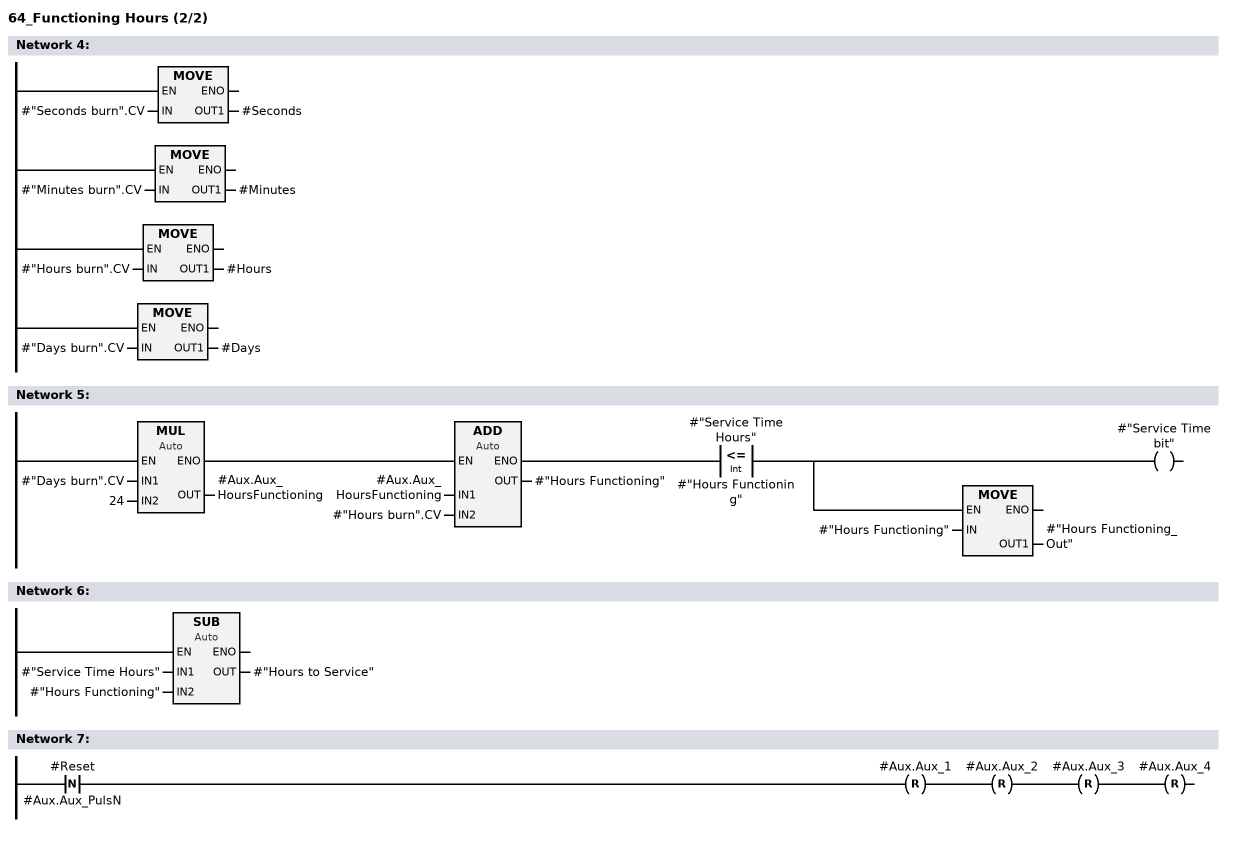
   RUNG wire#powerrail
      Move(in := #"Seconds burn".CV, out1 => #Seconds)
   END_RUNG
   RUNG wire#powerrail
      Move(in := #"Minutes burn".CV, out1 => #Minutes)
   END_RUNG
   RUNG wire#powerrail
      Move(in := #"Hours burn".CV, out1 => #Hours)
   END_RUNG
   RUNG wire#powerrail
      Move(in := #"Days burn".CV, out1 => #Days)
   END_RUNG
   // the same network as SCL:
   #Seconds := #"Seconds burn".CV;
   #Minutes := #"Minutes burn".CV;
   #Hours := #"Hours burn".CV;
   #Days := #"Days burn".CV;
END_REGION

REGION Network 5
   RUNG wire#powerrail
      Mul(in1 := #"Days burn".CV, in2 := 24, out => #Aux.Aux_HoursFunctioning)
      Add(in1 := #Aux.Aux_HoursFunctioning, in2 := #"Hours burn".CV, out => #"Hours Functioning")
      { S7_Templates := "SrcType := Int" } LE_Contact(in1 := #"Service Time Hours", in2 := #"Hours Functioning")
      wire#w1
      Coil( #"Service Time bit" )
   END_RUNG
   RUNG wire#w1
      Move(in := #"Hours Functioning", out1 => #"Hours Functioning_Out")
   END_RUNG
   // the same network as SCL:
   #Aux.Aux_HoursFunctioning := #"Days burn".CV * 24;
   #"Hours Functioning" := #Aux.Aux_HoursFunctioning + #"Hours burn".CV;
   #"Service Time bit" := #"Service Time Hours" <= #"Hours Functioning";
   IF #"Service Time bit" THEN #"Hours Functioning_Out" := #"Hours Functioning"; END_IF;
END_REGION

REGION Network 6
   RUNG wire#powerrail
      Sub(in1 := #"Service Time Hours", in2 := #"Hours Functioning", out => #"Hours to Service")
   END_RUNG
   // the same network as SCL:
   #"Hours to Service" := #"Service Time Hours" - #"Hours Functioning";
END_REGION

REGION Network 7
   RUNG wire#powerrail
      N_Contact(operand := #Reset, bit := #Aux.Aux_PulsN)
      R_Coil( #Aux.Aux_1 )
      R_Coil( #Aux.Aux_2 )
      R_Coil( #Aux.Aux_3 )
      R_Coil( #Aux.Aux_4 )
   END_RUNG
   // the same network as SCL:
   #_w1 := NOT #Reset AND #Aux.Aux_PulsN;   // falling edge of #Reset
   #Aux.Aux_PulsN := #Reset;
   IF #_w1 THEN
       #Aux.Aux_1 := FALSE;
       #Aux.Aux_2 := FALSE;
       #Aux.Aux_3 := FALSE;
       #Aux.Aux_4 := FALSE;
   END_IF;
END_REGION
END_FUNCTION_BLOCK

FUNCTION_BLOCK "503_ALARM CHCK II"   // FB507, LAD
{ S7_Optimized_Access := 'TRUE' }
VERSION : 0.1
   VAR_INPUT
      "Alarm Word 1" : Word;
      "Alarm Word Ack 1" : Word;
      "Alarm Word 2" : Word;
      "Alarm Word Ack 2" : Word;
      "Alarm Word 3" : Word;
      "Alarm Word Ack 3" : Word;
      "Alarm Word 4" : Word;
      "Alarm Word Ack 4" : Word;
      "Alarm Word 5" : Word;
      "Alarm Word Ack 5" : Word;
      "Alarm Word 6" : Word;
      "Alarm Word Ack 6" : Word;
      "Alarm Word 7" : Word;
      "Alarm Word Ack 7" : Word;
      "Alarm Word 8" : Word;
      "Alarm Word Ack 8" : Word;
      "Alarm Word 9" : Word;
      "Alarm Word 10" : Word;
      "Alarm Word 11" : Word;
      "Alarm Word 12" : Word;
      "Alarm Word 13" : Word;
      "Alarm Word 14" : Word;
      "Alarm Word 15" : Word;
      "Alarm Word 16" : Word;
      "Ack frequency" : Time;
      "Reset Alarm" : Bool;
   END_VAR
   VAR_OUTPUT
      Alarm : Bool;
      "New Alarm" : Bool;
      "Acknowledged Alarm" : Bool;
      Buzzer : Bool;
   END_VAR
   VAR
      "Alarm Word Interm 1" : Word;
      "Alarm Word Interm 2" : Word;
      "Alarm Word Interm 3" : Word;
      "Alarm Word Interm 4" : Word;
      "Alarm Word Interm 5" : Word;
      "Alarm Word Interm 6" : Word;
      "Alarm Word Interm 7" : Word;
      "Alarm Word Interm 8" : Word;
      "Alarm Word Interm 9" : Word;
      "Alarm Word Interm 10" : Word;
      "Alarm Word Interm 11" : Word;
      "Alarm Word Interm 12" : Word;
      "Alarm Word Interm 13" : Word;
      "Alarm Word Interm 14" : Word;
      "Alarm Word Interm 15" : Word;
      "Alarm Word Interm 16" : Word;
      "Alarm Word bool 1" : Bool;
      "Alarm Word bool 2" : Bool;
      "Alarm Word bool 3" : Bool;
      "Alarm Word bool 4" : Bool;
      "Alarm Word bool 5" : Bool;
      "Alarm Word bool 6" : Bool;
      "Alarm Word bool 7" : Bool;
      "Alarm Word bool 8" : Bool;
      "Alarm Word bool 9" : Bool;
      "Alarm Word bool 10" : Bool;
      "Alarm Word bool 11" : Bool;
      "Alarm Word bool 12" : Bool;
      "Alarm Word bool 13" : Bool;
      "Alarm Word bool 14" : Bool;
      "Alarm Word bool 15" : Bool;
      "Alarm Word bool 16" : Bool;
      True : Bool;
      False : Bool;
      "Delayed Alarm Reset" : TON_TIME;
      "Sound Alarm Delayed" : Bool;
      "SET TON" : TON_TIME;
      "RESET TON" : TON_TIME;
   END_VAR
   VAR_TEMP   // added for the SCL form of the ladder/FBD networks
      _w1 : Bool;
   END_VAR
BEGIN

REGION Network 1: True/False
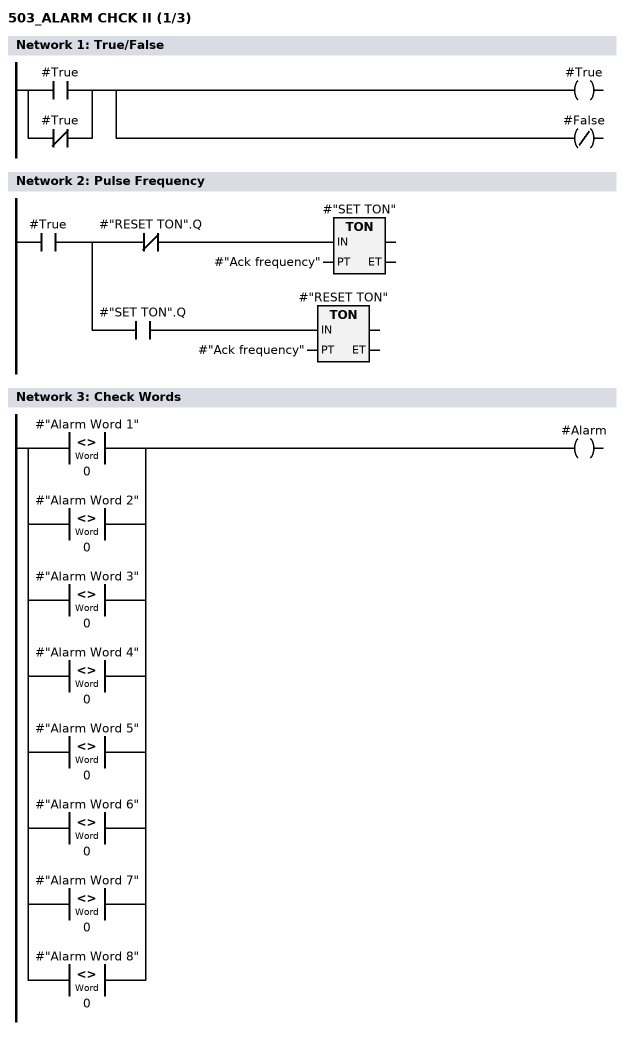
   RUNG wire#powerrail
      Contact( #True )
      wire#w1
      Coil( #True )
   END_RUNG
   RUNG wire#powerrail
      I_Contact( #True )
   END_RUNG wire#w1
   RUNG wire#w1
      I_Coil( #False )
   END_RUNG
   // the same network as SCL:
   #True := #True OR NOT #True;
   #False := NOT #True;
END_REGION

REGION Network 2: Pulse Frequency
   #"SET TON"(IN := #True AND NOT #"RESET TON".Q, PT := #"Ack frequency");   // TON
   #"RESET TON"(IN := #True AND #"SET TON".Q, PT := #"Ack frequency");   // TON
END_REGION

REGION Network 3: Check Words
   RUNG wire#powerrail
      { S7_Templates := "SrcType := Word" } NE_Contact(in1 := #"Alarm Word 1", in2 := 0)
      wire#w1
      Coil( #Alarm )
   END_RUNG
   RUNG wire#powerrail
      { S7_Templates := "SrcType := Word" } NE_Contact(in1 := #"Alarm Word 2", in2 := 0)
   END_RUNG wire#w1
   RUNG wire#powerrail
      { S7_Templates := "SrcType := Word" } NE_Contact(in1 := #"Alarm Word 3", in2 := 0)
   END_RUNG wire#w1
   RUNG wire#powerrail
      { S7_Templates := "SrcType := Word" } NE_Contact(in1 := #"Alarm Word 4", in2 := 0)
   END_RUNG wire#w1
   RUNG wire#powerrail
      { S7_Templates := "SrcType := Word" } NE_Contact(in1 := #"Alarm Word 5", in2 := 0)
   END_RUNG wire#w1
   RUNG wire#powerrail
      { S7_Templates := "SrcType := Word" } NE_Contact(in1 := #"Alarm Word 6", in2 := 0)
   END_RUNG wire#w1
   RUNG wire#powerrail
      { S7_Templates := "SrcType := Word" } NE_Contact(in1 := #"Alarm Word 7", in2 := 0)
   END_RUNG wire#w1
   RUNG wire#powerrail
      { S7_Templates := "SrcType := Word" } NE_Contact(in1 := #"Alarm Word 8", in2 := 0)
   END_RUNG wire#w1
   // the same network as SCL:
   #Alarm := (#"Alarm Word 1" <> 0) OR (#"Alarm Word 2" <> 0) OR (#"Alarm Word 3" <> 0) OR (#"Alarm Word 4" <> 0) OR (#"Alarm Word 5" <> 0) OR (#"Alarm Word 6" <> 0) OR (#"Alarm Word 7" <> 0) OR (#"Alarm Word 8" <> 0);
END_REGION

REGION Network 4: Check Words
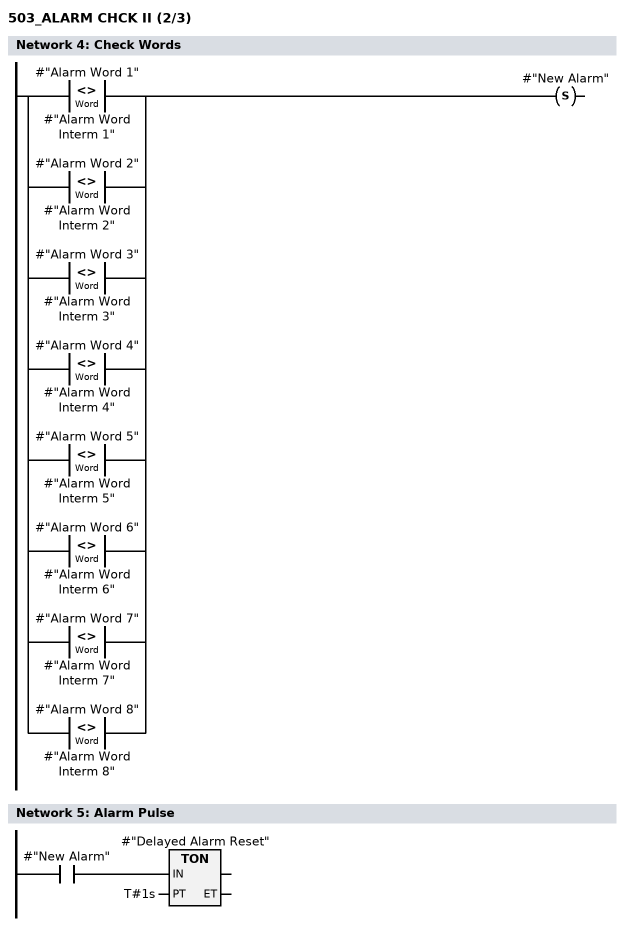
   RUNG wire#powerrail
      { S7_Templates := "SrcType := Word" } NE_Contact(in1 := #"Alarm Word 1", in2 := #"Alarm Word Interm 1")
      wire#w1
      S_Coil( #"New Alarm" )
   END_RUNG
   RUNG wire#powerrail
      { S7_Templates := "SrcType := Word" } NE_Contact(in1 := #"Alarm Word 2", in2 := #"Alarm Word Interm 2")
   END_RUNG wire#w1
   RUNG wire#powerrail
      { S7_Templates := "SrcType := Word" } NE_Contact(in1 := #"Alarm Word 3", in2 := #"Alarm Word Interm 3")
   END_RUNG wire#w1
   RUNG wire#powerrail
      { S7_Templates := "SrcType := Word" } NE_Contact(in1 := #"Alarm Word 4", in2 := #"Alarm Word Interm 4")
   END_RUNG wire#w1
   RUNG wire#powerrail
      { S7_Templates := "SrcType := Word" } NE_Contact(in1 := #"Alarm Word 5", in2 := #"Alarm Word Interm 5")
   END_RUNG wire#w1
   RUNG wire#powerrail
      { S7_Templates := "SrcType := Word" } NE_Contact(in1 := #"Alarm Word 6", in2 := #"Alarm Word Interm 6")
   END_RUNG wire#w1
   RUNG wire#powerrail
      { S7_Templates := "SrcType := Word" } NE_Contact(in1 := #"Alarm Word 7", in2 := #"Alarm Word Interm 7")
   END_RUNG wire#w1
   RUNG wire#powerrail
      { S7_Templates := "SrcType := Word" } NE_Contact(in1 := #"Alarm Word 8", in2 := #"Alarm Word Interm 8")
   END_RUNG wire#w1
   // the same network as SCL:
   IF (#"Alarm Word 1" <> #"Alarm Word Interm 1") OR (#"Alarm Word 2" <> #"Alarm Word Interm 2") OR (#"Alarm Word 3" <> #"Alarm Word Interm 3") OR (#"Alarm Word 4" <> #"Alarm Word Interm 4") OR (#"Alarm Word 5" <> #"Alarm Word Interm 5") OR (#"Alarm Word 6" <> #"Alarm Word Interm 6") OR (#"Alarm Word 7" <> #"Alarm Word Interm 7") OR (#"Alarm Word 8" <> #"Alarm Word Interm 8") THEN
       #"New Alarm" := TRUE;
   END_IF;
END_REGION

REGION Network 5: Alarm Pulse
   #"Delayed Alarm Reset"(IN := #"New Alarm", PT := T#1s);   // TON
END_REGION

REGION Network 6: Move Words
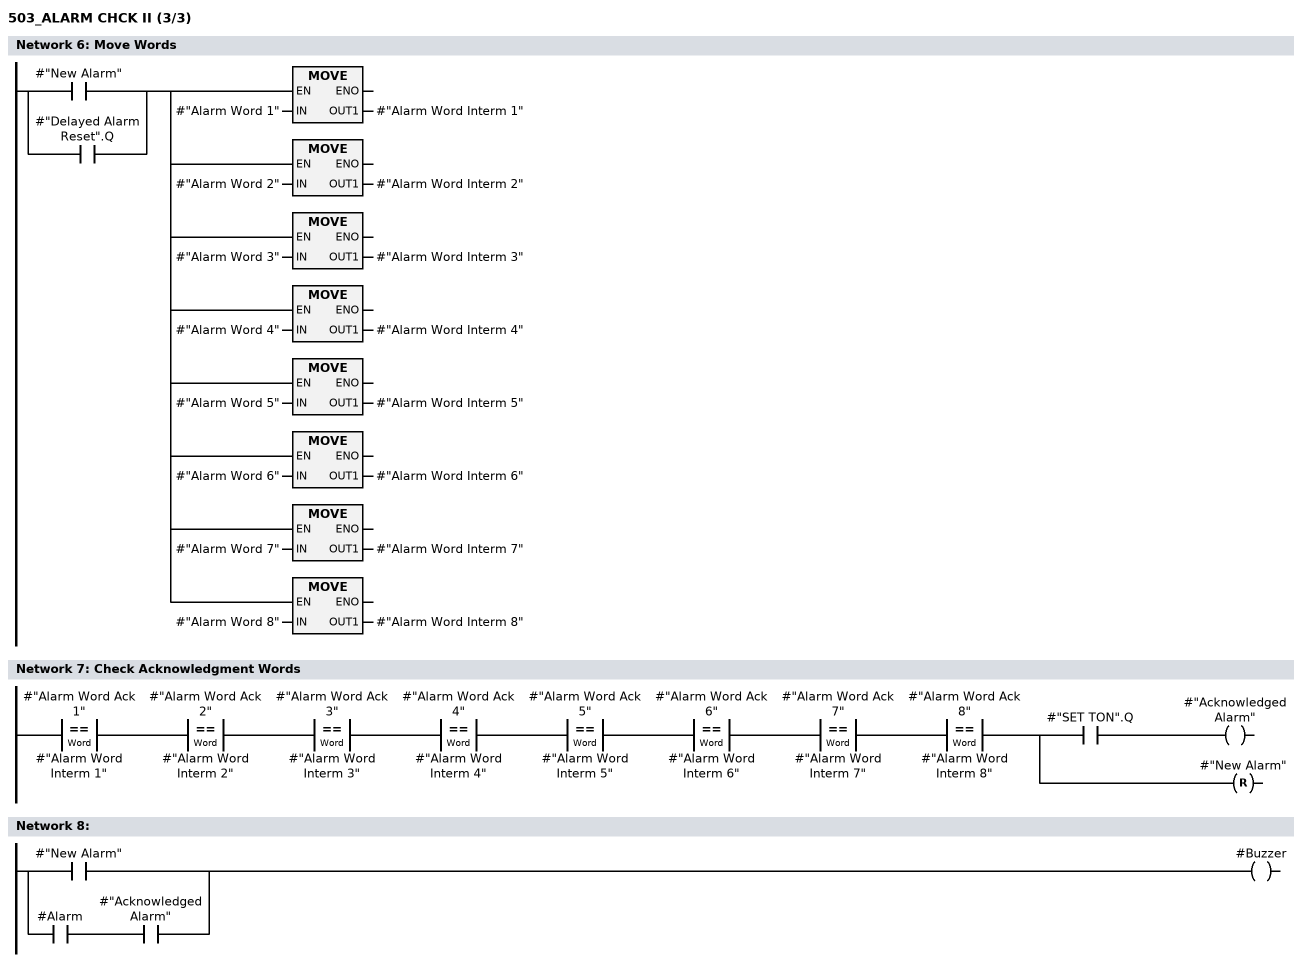
   RUNG wire#powerrail
      Contact( #"New Alarm" )
      wire#w1
      Move(in := #"Alarm Word 1", out1 => #"Alarm Word Interm 1")
   END_RUNG
   RUNG wire#powerrail
      Contact( #"Delayed Alarm Reset".Q )
   END_RUNG wire#w1
   RUNG wire#w1
      Move(in := #"Alarm Word 2", out1 => #"Alarm Word Interm 2")
   END_RUNG
   RUNG wire#w1
      Move(in := #"Alarm Word 3", out1 => #"Alarm Word Interm 3")
   END_RUNG
   RUNG wire#w1
      Move(in := #"Alarm Word 4", out1 => #"Alarm Word Interm 4")
   END_RUNG
   RUNG wire#w1
      Move(in := #"Alarm Word 5", out1 => #"Alarm Word Interm 5")
   END_RUNG
   RUNG wire#w1
      Move(in := #"Alarm Word 6", out1 => #"Alarm Word Interm 6")
   END_RUNG
   RUNG wire#w1
      Move(in := #"Alarm Word 7", out1 => #"Alarm Word Interm 7")
   END_RUNG
   RUNG wire#w1
      Move(in := #"Alarm Word 8", out1 => #"Alarm Word Interm 8")
   END_RUNG
   // the same network as SCL:
   IF #"New Alarm" OR #"Delayed Alarm Reset".Q THEN
       #"Alarm Word Interm 1" := #"Alarm Word 1";
       #"Alarm Word Interm 2" := #"Alarm Word 2";
       #"Alarm Word Interm 3" := #"Alarm Word 3";
       #"Alarm Word Interm 4" := #"Alarm Word 4";
       #"Alarm Word Interm 5" := #"Alarm Word 5";
       #"Alarm Word Interm 6" := #"Alarm Word 6";
       #"Alarm Word Interm 7" := #"Alarm Word 7";
       #"Alarm Word Interm 8" := #"Alarm Word 8";
   END_IF;
END_REGION

REGION Network 7: Check Acknowledgment Words
   RUNG wire#powerrail
      { S7_Templates := "SrcType := Word" } EQ_Contact(in1 := #"Alarm Word Ack 1", in2 := #"Alarm Word Interm 1")
      { S7_Templates := "SrcType := Word" } EQ_Contact(in1 := #"Alarm Word Ack 2", in2 := #"Alarm Word Interm 2")
      { S7_Templates := "SrcType := Word" } EQ_Contact(in1 := #"Alarm Word Ack 3", in2 := #"Alarm Word Interm 3")
      { S7_Templates := "SrcType := Word" } EQ_Contact(in1 := #"Alarm Word Ack 4", in2 := #"Alarm Word Interm 4")
      { S7_Templates := "SrcType := Word" } EQ_Contact(in1 := #"Alarm Word Ack 5", in2 := #"Alarm Word Interm 5")
      { S7_Templates := "SrcType := Word" } EQ_Contact(in1 := #"Alarm Word Ack 6", in2 := #"Alarm Word Interm 6")
      { S7_Templates := "SrcType := Word" } EQ_Contact(in1 := #"Alarm Word Ack 7", in2 := #"Alarm Word Interm 7")
      { S7_Templates := "SrcType := Word" } EQ_Contact(in1 := #"Alarm Word Ack 8", in2 := #"Alarm Word Interm 8")
      wire#w1
      Contact( #"SET TON".Q )
      Coil( #"Acknowledged Alarm" )
   END_RUNG
   RUNG wire#w1
      R_Coil( #"New Alarm" )
   END_RUNG
   // the same network as SCL:
   #_w1 := (#"Alarm Word Ack 1" = #"Alarm Word Interm 1") AND (#"Alarm Word Ack 2" = #"Alarm Word Interm 2") AND (#"Alarm Word Ack 3" = #"Alarm Word Interm 3") AND (#"Alarm Word Ack 4" = #"Alarm Word Interm 4") AND (#"Alarm Word Ack 5" = #"Alarm Word Interm 5") AND (#"Alarm Word Ack 6" = #"Alarm Word Interm 6") AND (#"Alarm Word Ack 7" = #"Alarm Word Interm 7") AND (#"Alarm Word Ack 8" = #"Alarm Word Interm 8");
   #"Acknowledged Alarm" := #_w1 AND #"SET TON".Q;
   IF #_w1 THEN #"New Alarm" := FALSE; END_IF;
END_REGION

REGION Network 8
   RUNG wire#powerrail
      Contact( #"New Alarm" )
      wire#w1
      Coil( #Buzzer )
   END_RUNG
   RUNG wire#powerrail
      Contact( #Alarm )
      Contact( #"Acknowledged Alarm" )
   END_RUNG wire#w1
   // the same network as SCL:
   #Buzzer := #"New Alarm" OR (#Alarm AND #"Acknowledged Alarm");
END_REGION
END_FUNCTION_BLOCK

FUNCTION_BLOCK "503_ALARM CHCK"   // FB508, LAD
{ S7_Optimized_Access := 'TRUE' }
VERSION : 0.1
   VAR_INPUT
      "Alarm Word 1" : Word;
      "Alarm Word 2" : Word;
      "Alarm Word 3" : Word;
      "Alarm Word 4" : Word;
      "Alarm Word 5" : Word;
      "Alarm Word 6" : Word;
      "Alarm Word 7" : Word;
      "Alarm Word 8" : Word;
      "Alarm Word 9" : Word;
      "Alarm Word 10" : Word;
      "Alarm Word 11" : Word;
      "Alarm Word 12" : Word;
      "Alarm Word 13" : Word;
      "Alarm Word 14" : Word;
      "Alarm Word 15" : Word;
      "Alarm Word 16" : Word;
      "Reset Alarm" : Bool;
   END_VAR
   VAR_OUTPUT
      "Sound Alarm" : Bool;
   END_VAR
   VAR
      "Alarm Word Interm 1" : Word;
      "Alarm Word Interm 2" : Word;
      "Alarm Word Interm 3" : Word;
      "Alarm Word Interm 4" : Word;
      "Alarm Word Interm 5" : Word;
      "Alarm Word Interm 6" : Word;
      "Alarm Word Interm 7" : Word;
      "Alarm Word Interm 8" : Word;
      "Alarm Word Interm 9" : Word;
      "Alarm Word Interm 10" : Word;
      "Alarm Word Interm 11" : Word;
      "Alarm Word Interm 12" : Word;
      "Alarm Word Interm 13" : Word;
      "Alarm Word Interm 14" : Word;
      "Alarm Word Interm 15" : Word;
      "Alarm Word Interm 16" : Word;
      "Alarm Word bool 1" : Bool;
      "Alarm Word bool 2" : Bool;
      "Alarm Word bool 3" : Bool;
      "Alarm Word bool 4" : Bool;
      "Alarm Word bool 5" : Bool;
      "Alarm Word bool 6" : Bool;
      "Alarm Word bool 7" : Bool;
      "Alarm Word bool 8" : Bool;
      "Alarm Word bool 9" : Bool;
      "Alarm Word bool 10" : Bool;
      "Alarm Word bool 11" : Bool;
      "Alarm Word bool 12" : Bool;
      "Alarm Word bool 13" : Bool;
      "Alarm Word bool 14" : Bool;
      "Alarm Word bool 15" : Bool;
      "Alarm Word bool 16" : Bool;
      "Delayed Alarm Reset" : TON_TIME;
   END_VAR
BEGIN

REGION Network 1: Check Words
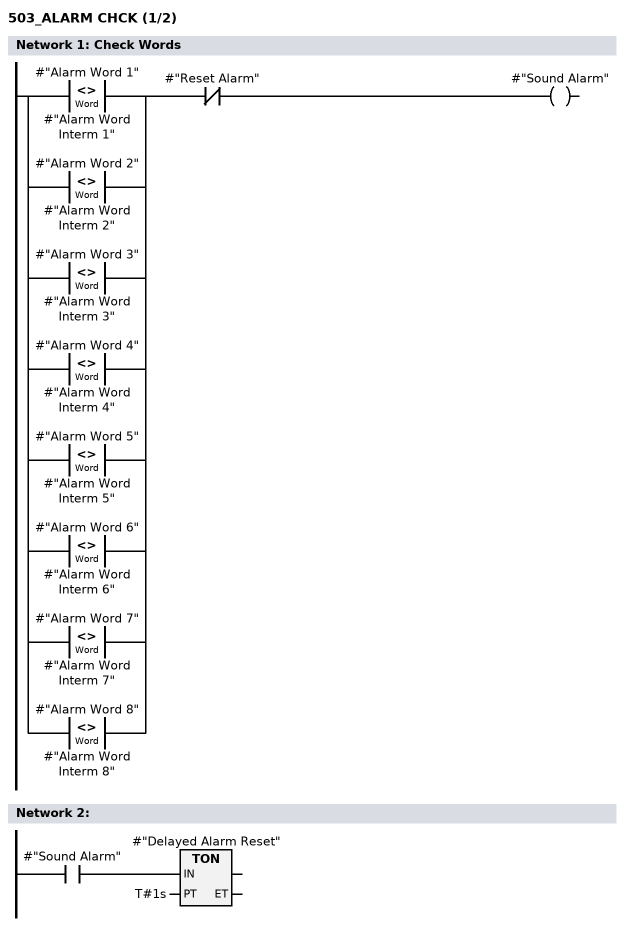
   RUNG wire#powerrail
      { S7_Templates := "SrcType := Word" } NE_Contact(in1 := #"Alarm Word 1", in2 := #"Alarm Word Interm 1")
      wire#w1
      I_Contact( #"Reset Alarm" )
      Coil( #"Sound Alarm" )
   END_RUNG
   RUNG wire#powerrail
      { S7_Templates := "SrcType := Word" } NE_Contact(in1 := #"Alarm Word 2", in2 := #"Alarm Word Interm 2")
   END_RUNG wire#w1
   RUNG wire#powerrail
      { S7_Templates := "SrcType := Word" } NE_Contact(in1 := #"Alarm Word 3", in2 := #"Alarm Word Interm 3")
   END_RUNG wire#w1
   RUNG wire#powerrail
      { S7_Templates := "SrcType := Word" } NE_Contact(in1 := #"Alarm Word 4", in2 := #"Alarm Word Interm 4")
   END_RUNG wire#w1
   RUNG wire#powerrail
      { S7_Templates := "SrcType := Word" } NE_Contact(in1 := #"Alarm Word 5", in2 := #"Alarm Word Interm 5")
   END_RUNG wire#w1
   RUNG wire#powerrail
      { S7_Templates := "SrcType := Word" } NE_Contact(in1 := #"Alarm Word 6", in2 := #"Alarm Word Interm 6")
   END_RUNG wire#w1
   RUNG wire#powerrail
      { S7_Templates := "SrcType := Word" } NE_Contact(in1 := #"Alarm Word 7", in2 := #"Alarm Word Interm 7")
   END_RUNG wire#w1
   RUNG wire#powerrail
      { S7_Templates := "SrcType := Word" } NE_Contact(in1 := #"Alarm Word 8", in2 := #"Alarm Word Interm 8")
   END_RUNG wire#w1
   // the same network as SCL:
   #"Sound Alarm" := ((#"Alarm Word 1" <> #"Alarm Word Interm 1") OR (#"Alarm Word 2" <> #"Alarm Word Interm 2") OR (#"Alarm Word 3" <> #"Alarm Word Interm 3") OR (#"Alarm Word 4" <> #"Alarm Word Interm 4") OR (#"Alarm Word 5" <> #"Alarm Word Interm 5") OR (#"Alarm Word 6" <> #"Alarm Word Interm 6") OR (#"Alarm Word 7" <> #"Alarm Word Interm 7") OR (#"Alarm Word 8" <> #"Alarm Word Interm 8")) AND NOT #"Reset Alarm";
END_REGION

REGION Network 2
   #"Delayed Alarm Reset"(IN := #"Sound Alarm", PT := T#1s);   // TON
END_REGION

REGION Network 3: Move Words
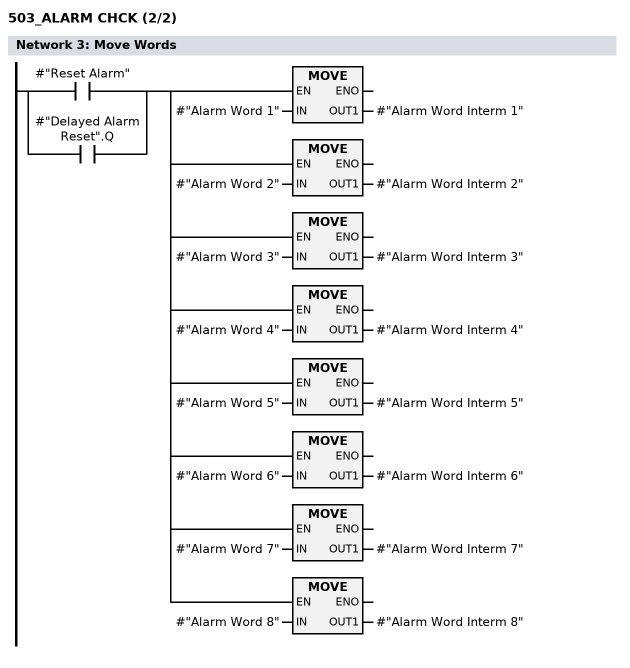
   RUNG wire#powerrail
      Contact( #"Reset Alarm" )
      wire#w1
      Move(in := #"Alarm Word 1", out1 => #"Alarm Word Interm 1")
   END_RUNG
   RUNG wire#powerrail
      Contact( #"Delayed Alarm Reset".Q )
   END_RUNG wire#w1
   RUNG wire#w1
      Move(in := #"Alarm Word 2", out1 => #"Alarm Word Interm 2")
   END_RUNG
   RUNG wire#w1
      Move(in := #"Alarm Word 3", out1 => #"Alarm Word Interm 3")
   END_RUNG
   RUNG wire#w1
      Move(in := #"Alarm Word 4", out1 => #"Alarm Word Interm 4")
   END_RUNG
   RUNG wire#w1
      Move(in := #"Alarm Word 5", out1 => #"Alarm Word Interm 5")
   END_RUNG
   RUNG wire#w1
      Move(in := #"Alarm Word 6", out1 => #"Alarm Word Interm 6")
   END_RUNG
   RUNG wire#w1
      Move(in := #"Alarm Word 7", out1 => #"Alarm Word Interm 7")
   END_RUNG
   RUNG wire#w1
      Move(in := #"Alarm Word 8", out1 => #"Alarm Word Interm 8")
   END_RUNG
   // the same network as SCL:
   IF #"Reset Alarm" OR #"Delayed Alarm Reset".Q THEN
       #"Alarm Word Interm 1" := #"Alarm Word 1";
       #"Alarm Word Interm 2" := #"Alarm Word 2";
       #"Alarm Word Interm 3" := #"Alarm Word 3";
       #"Alarm Word Interm 4" := #"Alarm Word 4";
       #"Alarm Word Interm 5" := #"Alarm Word 5";
       #"Alarm Word Interm 6" := #"Alarm Word 6";
       #"Alarm Word Interm 7" := #"Alarm Word 7";
       #"Alarm Word Interm 8" := #"Alarm Word 8";
   END_IF;
END_REGION
END_FUNCTION_BLOCK

FUNCTION_BLOCK "Evolving Setpoint"   // FB509, LAD
{ S7_Optimized_Access := 'TRUE' }
VERSION : 0.1
   VAR_INPUT
      Enable : Bool;
      Value : Real;
      Setpoint : Real;
      Gain : Real;
      Level_High : Real;
      Level_Low : Real;
   END_VAR
   VAR_OUTPUT
      Gain_Derived : Real;
      LevelBetter : Bool;
   END_VAR
   VAR
      "OFF Time" : TON_TIME;
      "On Time" : TON_TIME;
      Aux : Struct
         Aux_Derived : Bool;
         AuxSenzorDerivata1 : Real;
         AuxSenzorDerivata2 : Real;
         AuxSenzorDerivata11 : Real;
         AuxSenzorDerivata12 : Real;
         Puls_1 : Bool;
         Puls_2 : Bool;
         Puls_3 : Bool;
         Puls_4 : Bool;
         Gain_1 : Real;
      END_STRUCT;
      "Delay TOF" : TOF_TIME;
      "LevelBetter Delay" : TOF_TIME;
      "LevelBetter Prolong" : TOF_TIME;
   END_VAR
   VAR_TEMP   // added for the SCL form of the ladder/FBD networks
      _w1 : Bool;
      _w2 : Bool;
      _w3 : Bool;
      _w4 : Bool;
      _w5 : Bool;
      _w6 : Bool;
   END_VAR
BEGIN

REGION Network 1: Calcul derivata
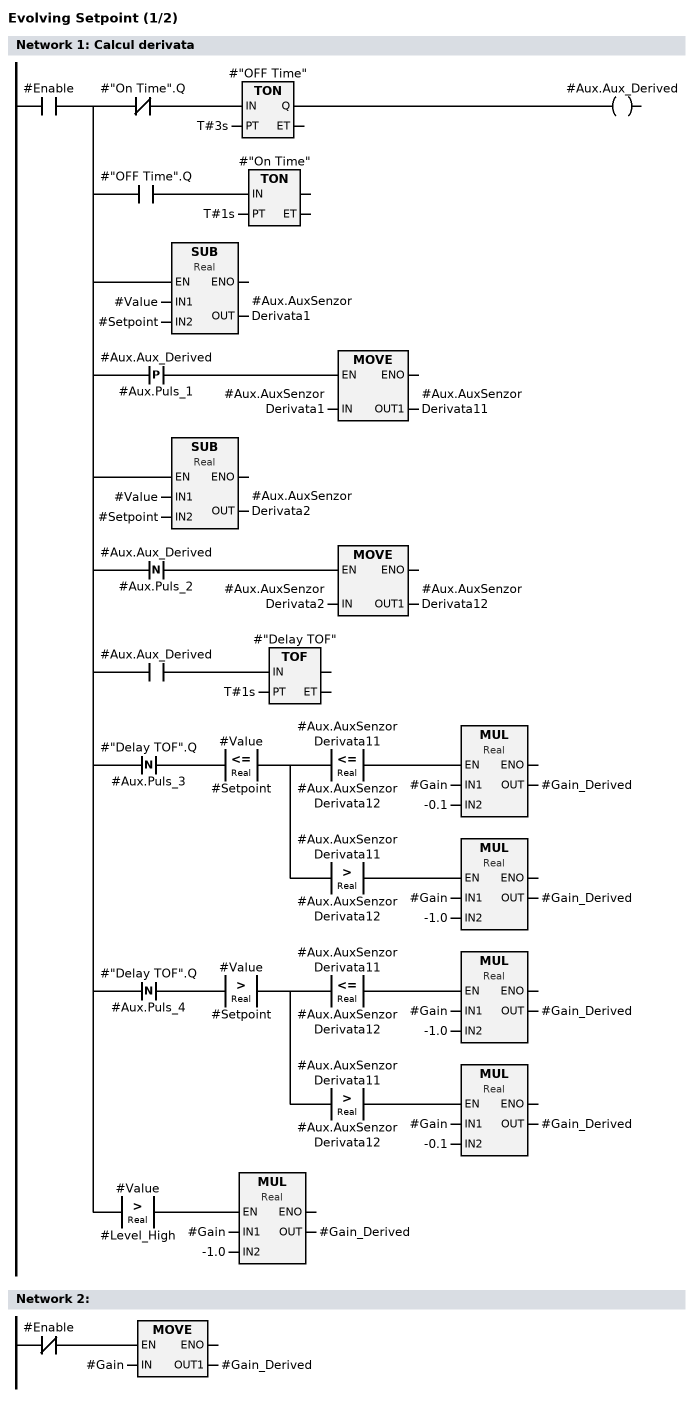
   #"OFF Time"(IN := #Enable AND NOT #"On Time".Q, PT := T#3s);   // TON
   #Aux.Aux_Derived := #"OFF Time".Q;
   #"On Time"(IN := #Enable AND #"OFF Time".Q, PT := T#1s);   // TON
   IF #Enable THEN #Aux.AuxSenzorDerivata1 := #Value - #Setpoint; END_IF;
   #_w1 := #Enable AND #Aux.Aux_Derived AND NOT #Aux.Puls_1;   // rising edge of #Aux.Aux_Derived
   #Aux.Puls_1 := #Aux.Aux_Derived;
   IF #_w1 THEN #Aux.AuxSenzorDerivata11 := #Aux.AuxSenzorDerivata1; END_IF;
   IF #Enable THEN #Aux.AuxSenzorDerivata2 := #Value - #Setpoint; END_IF;
   #_w2 := #Enable AND NOT #Aux.Aux_Derived AND #Aux.Puls_2;   // falling edge of #Aux.Aux_Derived
   #Aux.Puls_2 := #Aux.Aux_Derived;
   IF #_w2 THEN #Aux.AuxSenzorDerivata12 := #Aux.AuxSenzorDerivata2; END_IF;
   #"Delay TOF"(IN := #Enable AND #Aux.Aux_Derived, PT := T#1s);   // TOF
   #_w3 := #Enable AND NOT #"Delay TOF".Q AND #Aux.Puls_3;   // falling edge of #"Delay TOF".Q
   #Aux.Puls_3 := #"Delay TOF".Q;
   #_w4 := #_w3 AND (#Value <= #Setpoint);
   IF #_w4 AND (#Aux.AuxSenzorDerivata11 <= #Aux.AuxSenzorDerivata12) THEN
       #Gain_Derived := #Gain * (-0.1);
   END_IF;
   IF #_w4 AND (#Aux.AuxSenzorDerivata11 > #Aux.AuxSenzorDerivata12) THEN
       #Gain_Derived := #Gain * (-1.0);
   END_IF;
   #_w5 := #Enable AND NOT #"Delay TOF".Q AND #Aux.Puls_4;   // falling edge of #"Delay TOF".Q
   #Aux.Puls_4 := #"Delay TOF".Q;
   #_w6 := #_w5 AND (#Value > #Setpoint);
   IF #_w6 AND (#Aux.AuxSenzorDerivata11 <= #Aux.AuxSenzorDerivata12) THEN
       #Gain_Derived := #Gain * (-1.0);
   END_IF;
   IF #_w6 AND (#Aux.AuxSenzorDerivata11 > #Aux.AuxSenzorDerivata12) THEN
       #Gain_Derived := #Gain * (-0.1);
   END_IF;
   IF #Enable AND (#Value > #Level_High) THEN #Gain_Derived := #Gain * (-1.0); END_IF;
END_REGION

REGION Network 2
   RUNG wire#powerrail
      I_Contact( #Enable )
      { S7_GenerateENO := "TRUE" } Move(in := #Gain, out1 => #Gain_Derived)
   END_RUNG
   // the same network as SCL:
   IF NOT #Enable THEN #Gain_Derived := #Gain; END_IF;
END_REGION

REGION Network 3: Neautorizare pompa la imbunatatirea nivelului
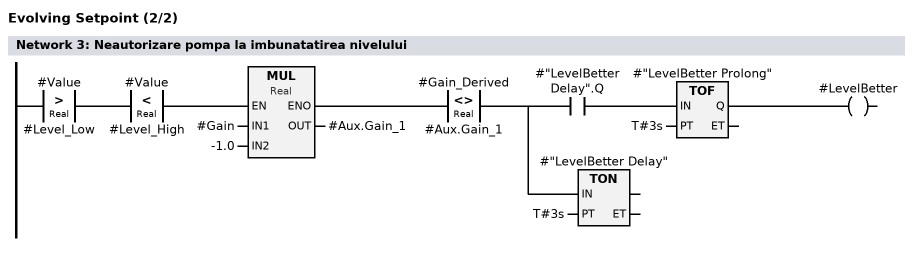
   // ENO of a box is taken as its EN; it also drops when the box reports an error
   #_w1 := (#Value > #Level_Low) AND (#Value < #Level_High);
   IF #_w1 THEN #Aux.Gain_1 := #Gain * (-1.0); END_IF;
   #_w2 := #_w1 AND (#Gain_Derived <> #Aux.Gain_1);
   #"LevelBetter Prolong"(IN := #_w2 AND #"LevelBetter Delay".Q, PT := T#3s);   // TOF
   #LevelBetter := #"LevelBetter Prolong".Q;
   #"LevelBetter Delay"(IN := #_w2, PT := T#3s);   // TON
END_REGION
END_FUNCTION_BLOCK

FUNCTION_BLOCK "Animation"   // FB515, LAD
{ S7_Optimized_Access := 'TRUE' }
VERSION : 0.1
   VAR_INPUT
      Run : Bool;
      Revert : Bool := true;
      "States Number" : Int := 10;
      Period : Time := T#250ms;
   END_VAR
   VAR_OUTPUT
      Animation : Int;
   END_VAR
   VAR RETAIN
      "Animation State" : CTU_INT;
      Reset : Bool;
   END_VAR
   VAR
      "Revert Aux" : Bool;
      LD : Bool;
      OFF : TON_TIME;
      ON : TON_TIME;
   END_VAR
BEGIN

REGION Network 1